(* Logix 5000 project; controller FV vendor 1 type 14 code 217 rev 31.11; software revision 31.00; part 20 of 63 *)
(* tags used below, declared in another part *)
   CheckTimeMask : INT;
   Delphi_Does_Eng_Func : BOOL;
   FR_FV26_AV04 : PlantItem;   // FV26_AV04
   FR_FV26_AV05 : PlantItem;   // FV26_AV05
   FR_FV26_AV06 : PlantItem;   // FV26_AV06
   FR_FV26_AV07 : PlantItem;   // FV26_AV07
   FR_FV27_AV01 : PlantItem;   // FV27_AV01
   FR_FV27_AV04 : PlantItem;   // FV27_AV04
   FR_FV27_AV05 : PlantItem;   // FV27_AV05
   FR_FV27_AV06 : PlantItem;   // FV27_AV06
   FR_FV27_AV07 : PlantItem;   // FV27_AV07
   FR_N255 : INT[265];   // CHECKWORDS
   FR_VB1_AV01 : PlantItem;   // VB1_AV01
   FR_VB1_AV02 : PlantItem;   // VB1_AV02
   FR_VB1_AV03 : PlantItem;   // VB1_AV03
   FR_VB1_AV04 : PlantItem;   // VB1_AV04
   TempChecktime : DINT;
(* FR_Common, continued *)

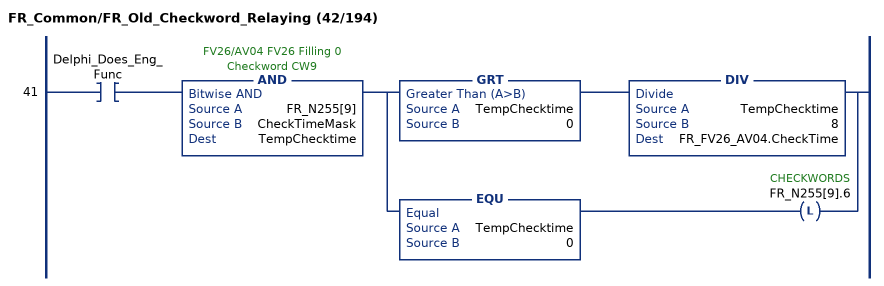
   [picture p346: FR_Common/FR_Old_Checkword_Relaying rungs 41-41]
   41: XIC(Delphi_Does_Eng_Func)AND(FR_N255[9],CheckTimeMask,TempChecktime)[GRT(TempChecktime,0) DIV(TempChecktime,8,FR_FV26_AV04.CheckTime) ,EQU(TempChecktime,0) OTL(FR_N255[9].6) ];
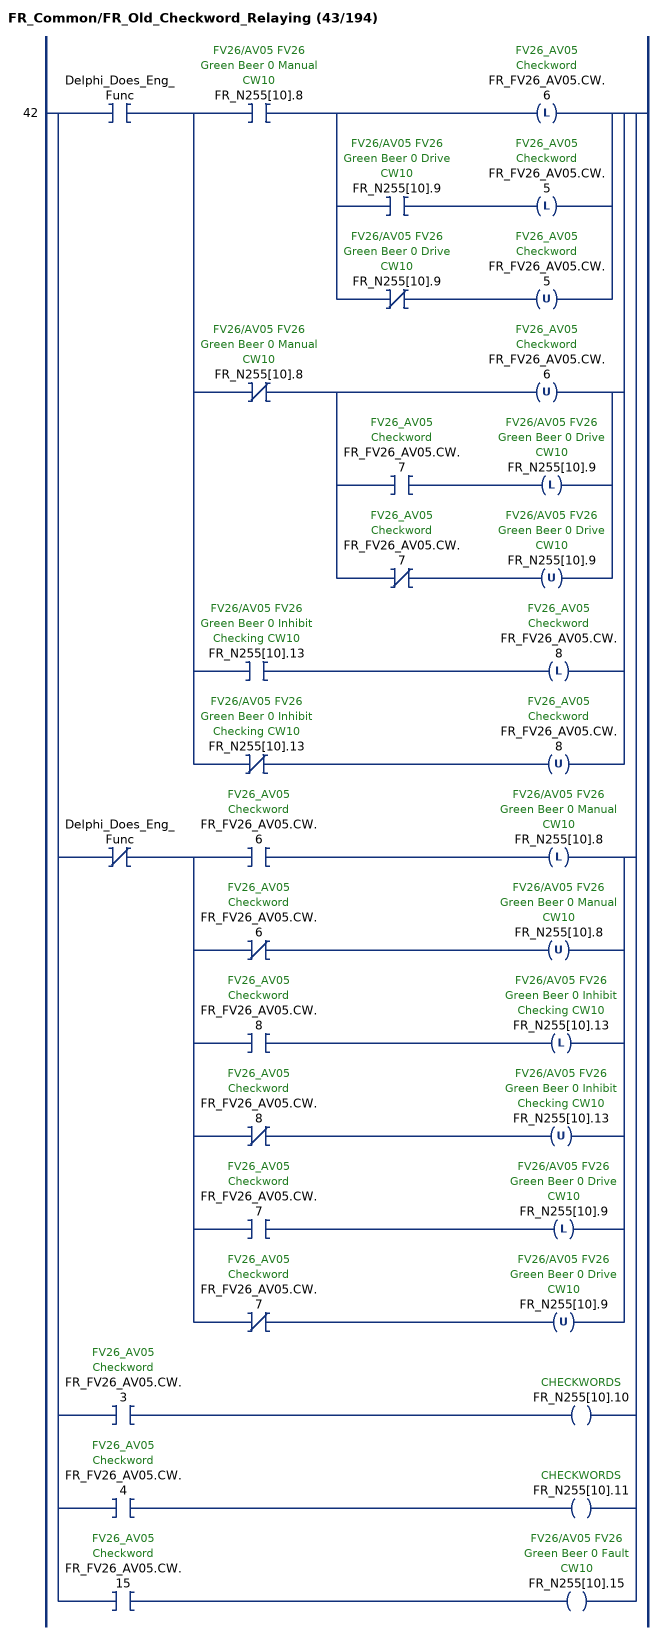
   42: [XIC(Delphi_Does_Eng_Func) [[XIC(FR_N255[10].8) [OTL(FR_FV26_AV05.CW.6) ,XIC(FR_N255[10].9) OTL(FR_FV26_AV05.CW.5) ,XIO(FR_N255[10].9) OTU(FR_FV26_AV05.CW.5) ] ,XIO(FR_N255[10].8) [OTU(FR_FV26_AV05.CW.6) ,[XIC(FR_FV26_AV05.CW.7) OTL(FR_N255[10].9) ,XIO(FR_FV26_AV05.CW.7) OTU(FR_N255[10].9) ] ] ] ,[XIC(FR_N255[10].13) OTL(FR_FV26_AV05.CW.8) ,XIO(FR_N255[10].13) OTU(FR_FV26_AV05.CW.8) ] ] ,XIO(Delphi_Does_Eng_Func) [[XIC(FR_FV26_AV05.CW.6) OTL(FR_N255[10].8) ,XIO(FR_FV26_AV05.CW.6) OTU(FR_N255[10].8) ] ,[XIC(FR_FV26_AV05.CW.8) OTL(FR_N255[10].13) ,XIO(FR_FV26_AV05.CW.8) OTU(FR_N255[10].13) ] ,[XIC(FR_FV26_AV05.CW.7) OTL(FR_N255[10].9) ,XIO(FR_FV26_AV05.CW.7) OTU(FR_N255[10].9) ] ] ,XIC(FR_FV26_AV05.CW.3) OTE(FR_N255[10].10) ,XIC(FR_FV26_AV05.CW.4) OTE(FR_N255[10].11) ,XIC(FR_FV26_AV05.CW.15) OTE(FR_N255[10].15) ];
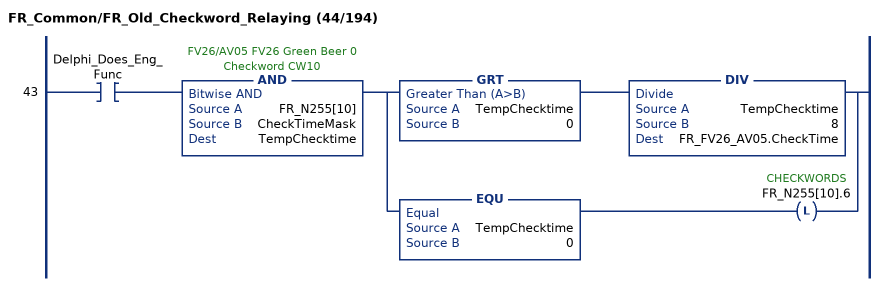
   43: XIC(Delphi_Does_Eng_Func)AND(FR_N255[10],CheckTimeMask,TempChecktime)[GRT(TempChecktime,0) DIV(TempChecktime,8,FR_FV26_AV05.CheckTime) ,EQU(TempChecktime,0) OTL(FR_N255[10].6) ];
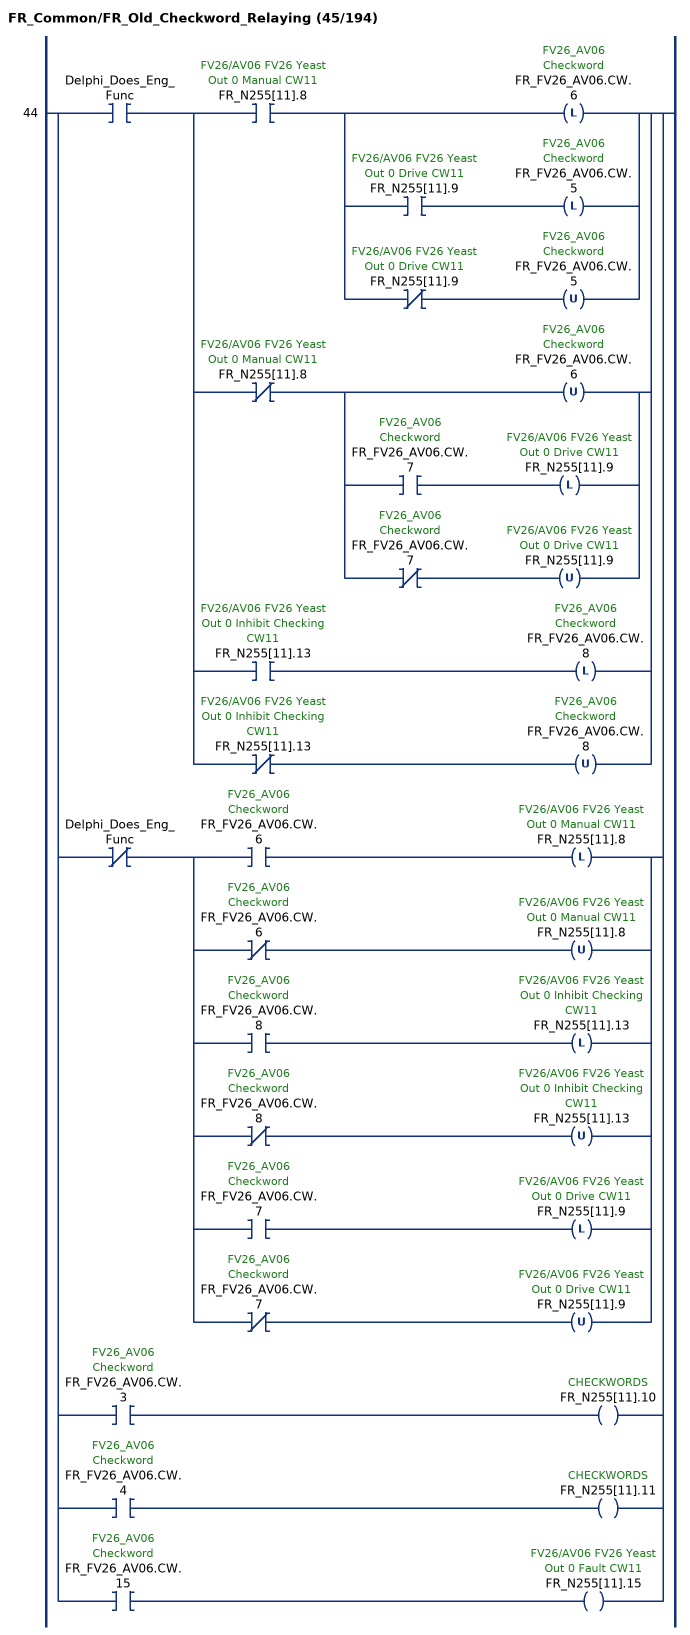
   44: [XIC(Delphi_Does_Eng_Func) [[XIC(FR_N255[11].8) [OTL(FR_FV26_AV06.CW.6) ,XIC(FR_N255[11].9) OTL(FR_FV26_AV06.CW.5) ,XIO(FR_N255[11].9) OTU(FR_FV26_AV06.CW.5) ] ,XIO(FR_N255[11].8) [OTU(FR_FV26_AV06.CW.6) ,[XIC(FR_FV26_AV06.CW.7) OTL(FR_N255[11].9) ,XIO(FR_FV26_AV06.CW.7) OTU(FR_N255[11].9) ] ] ] ,[XIC(FR_N255[11].13) OTL(FR_FV26_AV06.CW.8) ,XIO(FR_N255[11].13) OTU(FR_FV26_AV06.CW.8) ] ] ,XIO(Delphi_Does_Eng_Func) [[XIC(FR_FV26_AV06.CW.6) OTL(FR_N255[11].8) ,XIO(FR_FV26_AV06.CW.6) OTU(FR_N255[11].8) ] ,[XIC(FR_FV26_AV06.CW.8) OTL(FR_N255[11].13) ,XIO(FR_FV26_AV06.CW.8) OTU(FR_N255[11].13) ] ,[XIC(FR_FV26_AV06.CW.7) OTL(FR_N255[11].9) ,XIO(FR_FV26_AV06.CW.7) OTU(FR_N255[11].9) ] ] ,XIC(FR_FV26_AV06.CW.3) OTE(FR_N255[11].10) ,XIC(FR_FV26_AV06.CW.4) OTE(FR_N255[11].11) ,XIC(FR_FV26_AV06.CW.15) OTE(FR_N255[11].15) ];
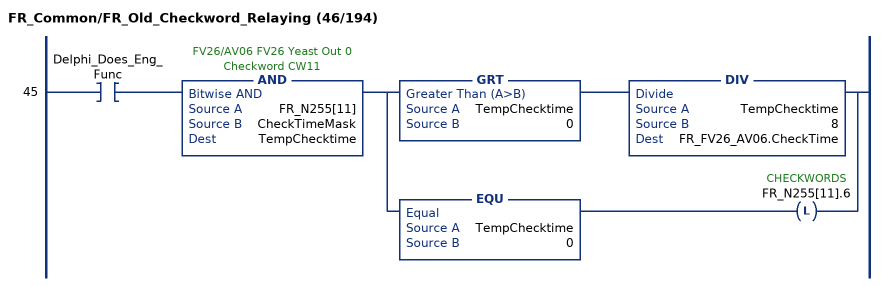
   45: XIC(Delphi_Does_Eng_Func)AND(FR_N255[11],CheckTimeMask,TempChecktime)[GRT(TempChecktime,0) DIV(TempChecktime,8,FR_FV26_AV06.CheckTime) ,EQU(TempChecktime,0) OTL(FR_N255[11].6) ];
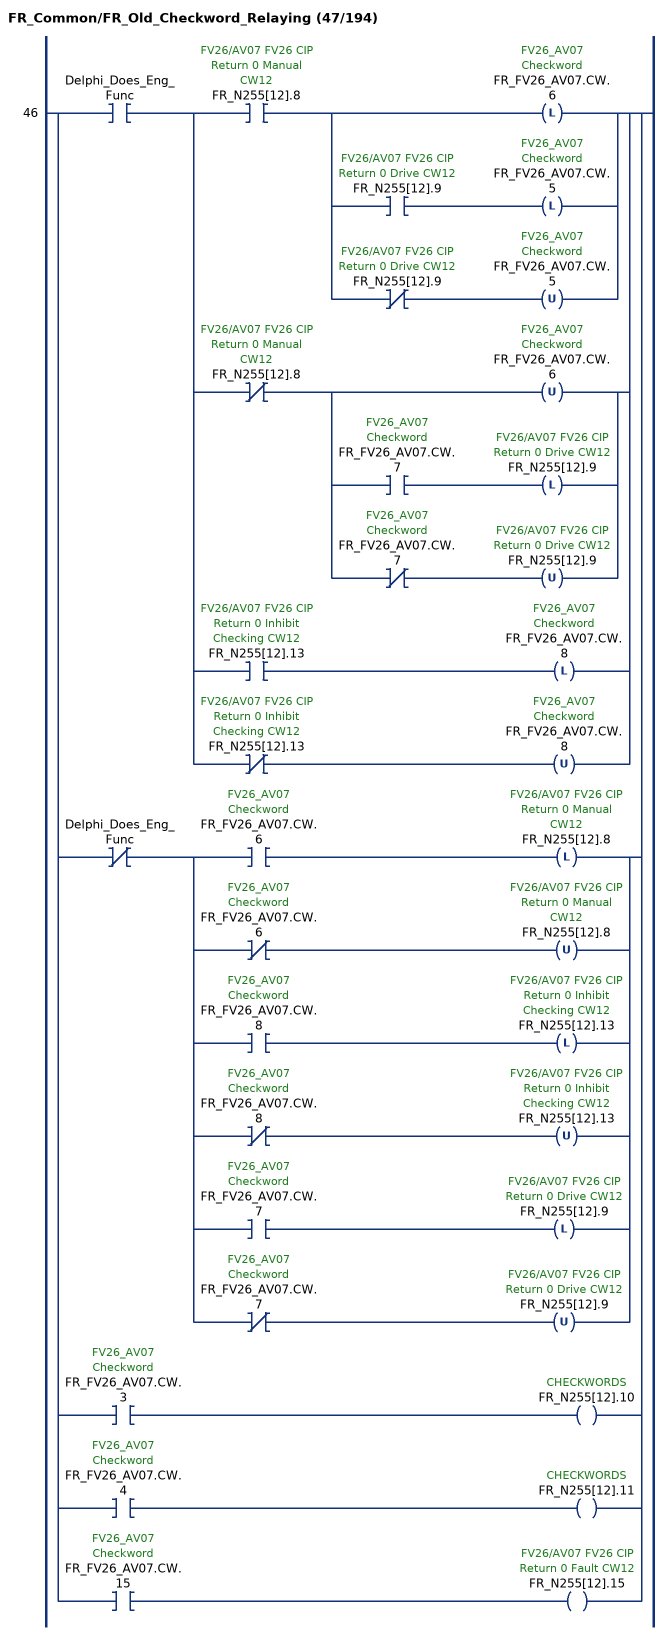
   46: [XIC(Delphi_Does_Eng_Func) [[XIC(FR_N255[12].8) [OTL(FR_FV26_AV07.CW.6) ,XIC(FR_N255[12].9) OTL(FR_FV26_AV07.CW.5) ,XIO(FR_N255[12].9) OTU(FR_FV26_AV07.CW.5) ] ,XIO(FR_N255[12].8) [OTU(FR_FV26_AV07.CW.6) ,[XIC(FR_FV26_AV07.CW.7) OTL(FR_N255[12].9) ,XIO(FR_FV26_AV07.CW.7) OTU(FR_N255[12].9) ] ] ] ,[XIC(FR_N255[12].13) OTL(FR_FV26_AV07.CW.8) ,XIO(FR_N255[12].13) OTU(FR_FV26_AV07.CW.8) ] ] ,XIO(Delphi_Does_Eng_Func) [[XIC(FR_FV26_AV07.CW.6) OTL(FR_N255[12].8) ,XIO(FR_FV26_AV07.CW.6) OTU(FR_N255[12].8) ] ,[XIC(FR_FV26_AV07.CW.8) OTL(FR_N255[12].13) ,XIO(FR_FV26_AV07.CW.8) OTU(FR_N255[12].13) ] ,[XIC(FR_FV26_AV07.CW.7) OTL(FR_N255[12].9) ,XIO(FR_FV26_AV07.CW.7) OTU(FR_N255[12].9) ] ] ,XIC(FR_FV26_AV07.CW.3) OTE(FR_N255[12].10) ,XIC(FR_FV26_AV07.CW.4) OTE(FR_N255[12].11) ,XIC(FR_FV26_AV07.CW.15) OTE(FR_N255[12].15) ];
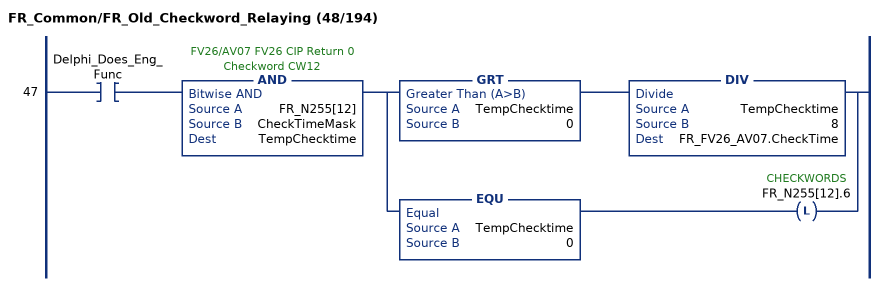
   47: XIC(Delphi_Does_Eng_Func)AND(FR_N255[12],CheckTimeMask,TempChecktime)[GRT(TempChecktime,0) DIV(TempChecktime,8,FR_FV26_AV07.CheckTime) ,EQU(TempChecktime,0) OTL(FR_N255[12].6) ];
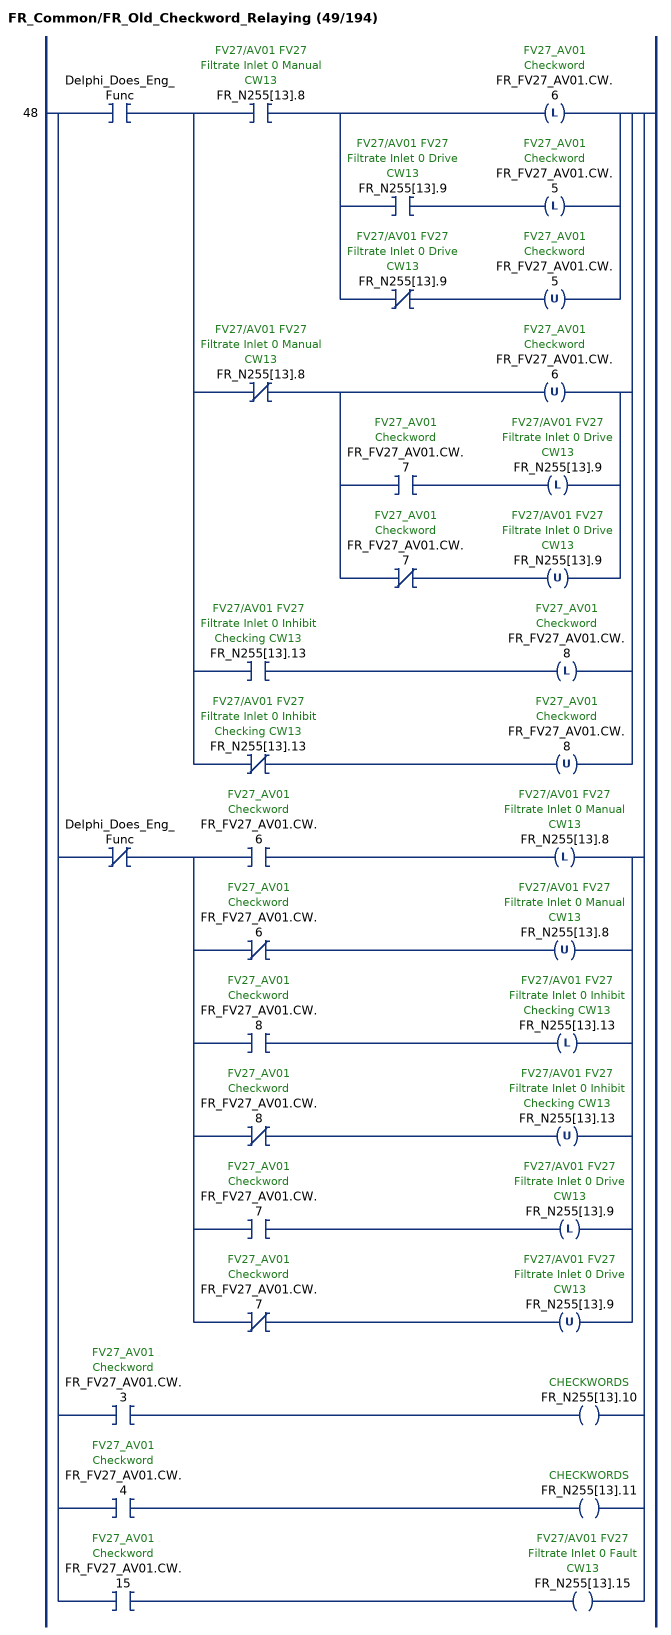
   48: [XIC(Delphi_Does_Eng_Func) [[XIC(FR_N255[13].8) [OTL(FR_FV27_AV01.CW.6) ,XIC(FR_N255[13].9) OTL(FR_FV27_AV01.CW.5) ,XIO(FR_N255[13].9) OTU(FR_FV27_AV01.CW.5) ] ,XIO(FR_N255[13].8) [OTU(FR_FV27_AV01.CW.6) ,[XIC(FR_FV27_AV01.CW.7) OTL(FR_N255[13].9) ,XIO(FR_FV27_AV01.CW.7) OTU(FR_N255[13].9) ] ] ] ,[XIC(FR_N255[13].13) OTL(FR_FV27_AV01.CW.8) ,XIO(FR_N255[13].13) OTU(FR_FV27_AV01.CW.8) ] ] ,XIO(Delphi_Does_Eng_Func) [[XIC(FR_FV27_AV01.CW.6) OTL(FR_N255[13].8) ,XIO(FR_FV27_AV01.CW.6) OTU(FR_N255[13].8) ] ,[XIC(FR_FV27_AV01.CW.8) OTL(FR_N255[13].13) ,XIO(FR_FV27_AV01.CW.8) OTU(FR_N255[13].13) ] ,[XIC(FR_FV27_AV01.CW.7) OTL(FR_N255[13].9) ,XIO(FR_FV27_AV01.CW.7) OTU(FR_N255[13].9) ] ] ,XIC(FR_FV27_AV01.CW.3) OTE(FR_N255[13].10) ,XIC(FR_FV27_AV01.CW.4) OTE(FR_N255[13].11) ,XIC(FR_FV27_AV01.CW.15) OTE(FR_N255[13].15) ];
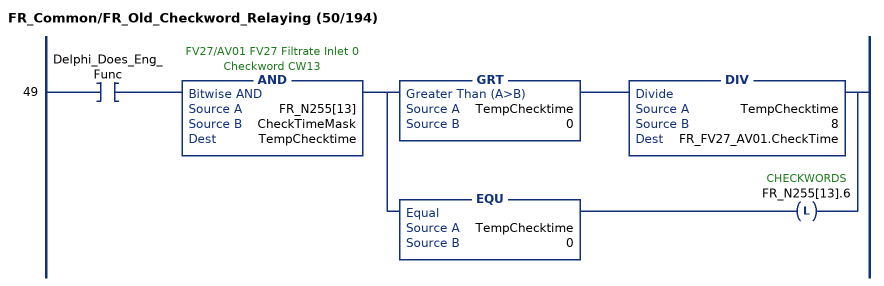
   49: XIC(Delphi_Does_Eng_Func)AND(FR_N255[13],CheckTimeMask,TempChecktime)[GRT(TempChecktime,0) DIV(TempChecktime,8,FR_FV27_AV01.CheckTime) ,EQU(TempChecktime,0) OTL(FR_N255[13].6) ];
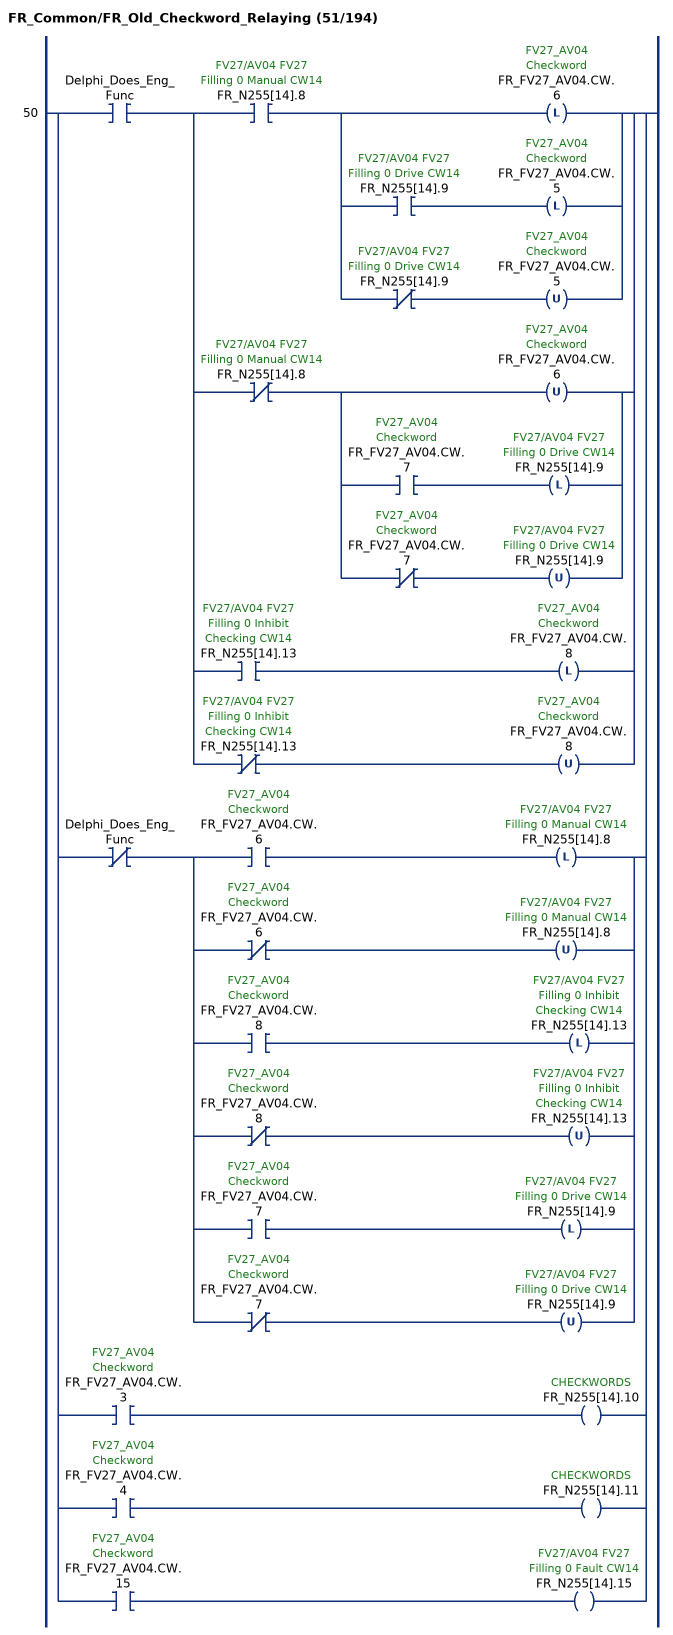
   50: [XIC(Delphi_Does_Eng_Func) [[XIC(FR_N255[14].8) [OTL(FR_FV27_AV04.CW.6) ,XIC(FR_N255[14].9) OTL(FR_FV27_AV04.CW.5) ,XIO(FR_N255[14].9) OTU(FR_FV27_AV04.CW.5) ] ,XIO(FR_N255[14].8) [OTU(FR_FV27_AV04.CW.6) ,[XIC(FR_FV27_AV04.CW.7) OTL(FR_N255[14].9) ,XIO(FR_FV27_AV04.CW.7) OTU(FR_N255[14].9) ] ] ] ,[XIC(FR_N255[14].13) OTL(FR_FV27_AV04.CW.8) ,XIO(FR_N255[14].13) OTU(FR_FV27_AV04.CW.8) ] ] ,XIO(Delphi_Does_Eng_Func) [[XIC(FR_FV27_AV04.CW.6) OTL(FR_N255[14].8) ,XIO(FR_FV27_AV04.CW.6) OTU(FR_N255[14].8) ] ,[XIC(FR_FV27_AV04.CW.8) OTL(FR_N255[14].13) ,XIO(FR_FV27_AV04.CW.8) OTU(FR_N255[14].13) ] ,[XIC(FR_FV27_AV04.CW.7) OTL(FR_N255[14].9) ,XIO(FR_FV27_AV04.CW.7) OTU(FR_N255[14].9) ] ] ,XIC(FR_FV27_AV04.CW.3) OTE(FR_N255[14].10) ,XIC(FR_FV27_AV04.CW.4) OTE(FR_N255[14].11) ,XIC(FR_FV27_AV04.CW.15) OTE(FR_N255[14].15) ];
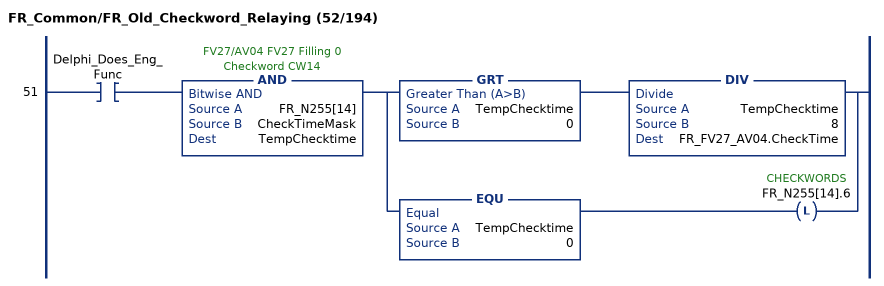
   51: XIC(Delphi_Does_Eng_Func)AND(FR_N255[14],CheckTimeMask,TempChecktime)[GRT(TempChecktime,0) DIV(TempChecktime,8,FR_FV27_AV04.CheckTime) ,EQU(TempChecktime,0) OTL(FR_N255[14].6) ];
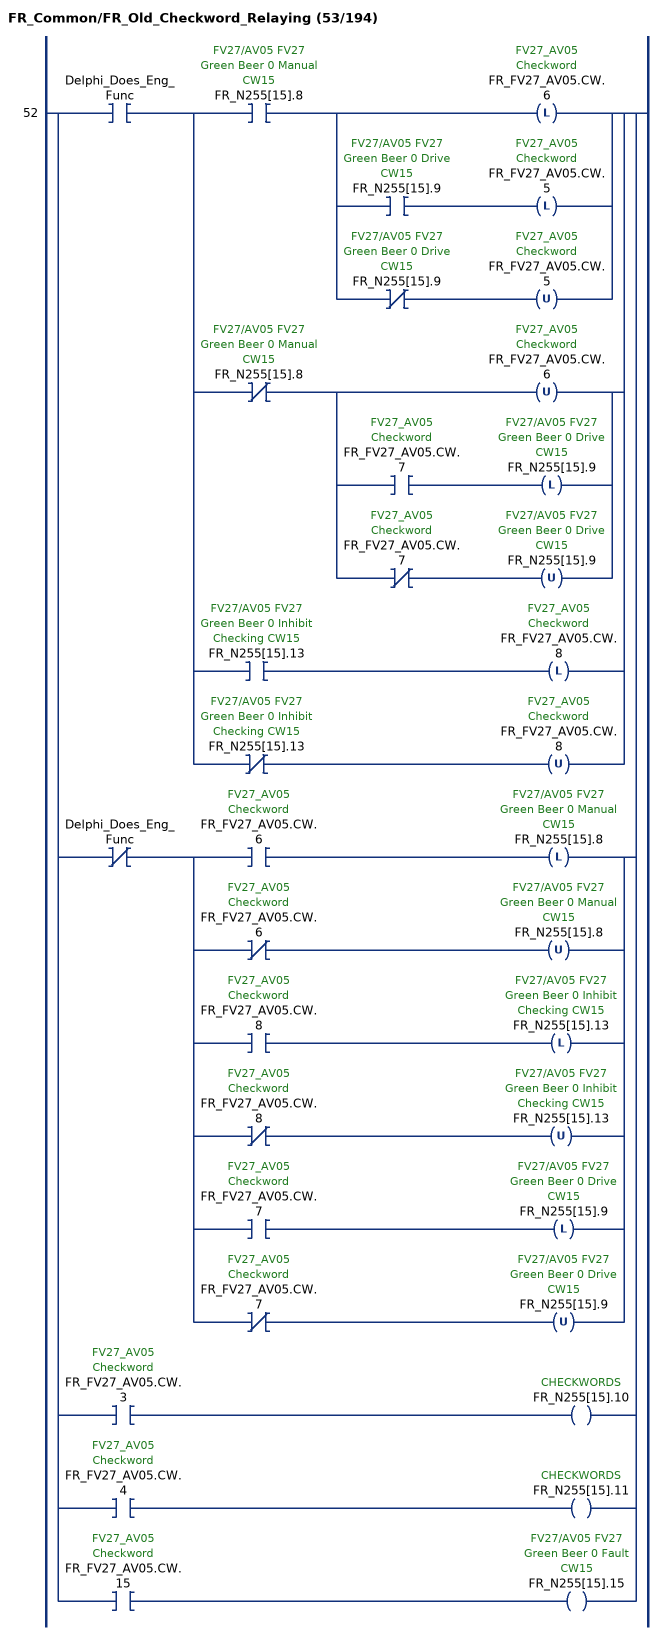
   52: [XIC(Delphi_Does_Eng_Func) [[XIC(FR_N255[15].8) [OTL(FR_FV27_AV05.CW.6) ,XIC(FR_N255[15].9) OTL(FR_FV27_AV05.CW.5) ,XIO(FR_N255[15].9) OTU(FR_FV27_AV05.CW.5) ] ,XIO(FR_N255[15].8) [OTU(FR_FV27_AV05.CW.6) ,[XIC(FR_FV27_AV05.CW.7) OTL(FR_N255[15].9) ,XIO(FR_FV27_AV05.CW.7) OTU(FR_N255[15].9) ] ] ] ,[XIC(FR_N255[15].13) OTL(FR_FV27_AV05.CW.8) ,XIO(FR_N255[15].13) OTU(FR_FV27_AV05.CW.8) ] ] ,XIO(Delphi_Does_Eng_Func) [[XIC(FR_FV27_AV05.CW.6) OTL(FR_N255[15].8) ,XIO(FR_FV27_AV05.CW.6) OTU(FR_N255[15].8) ] ,[XIC(FR_FV27_AV05.CW.8) OTL(FR_N255[15].13) ,XIO(FR_FV27_AV05.CW.8) OTU(FR_N255[15].13) ] ,[XIC(FR_FV27_AV05.CW.7) OTL(FR_N255[15].9) ,XIO(FR_FV27_AV05.CW.7) OTU(FR_N255[15].9) ] ] ,XIC(FR_FV27_AV05.CW.3) OTE(FR_N255[15].10) ,XIC(FR_FV27_AV05.CW.4) OTE(FR_N255[15].11) ,XIC(FR_FV27_AV05.CW.15) OTE(FR_N255[15].15) ];